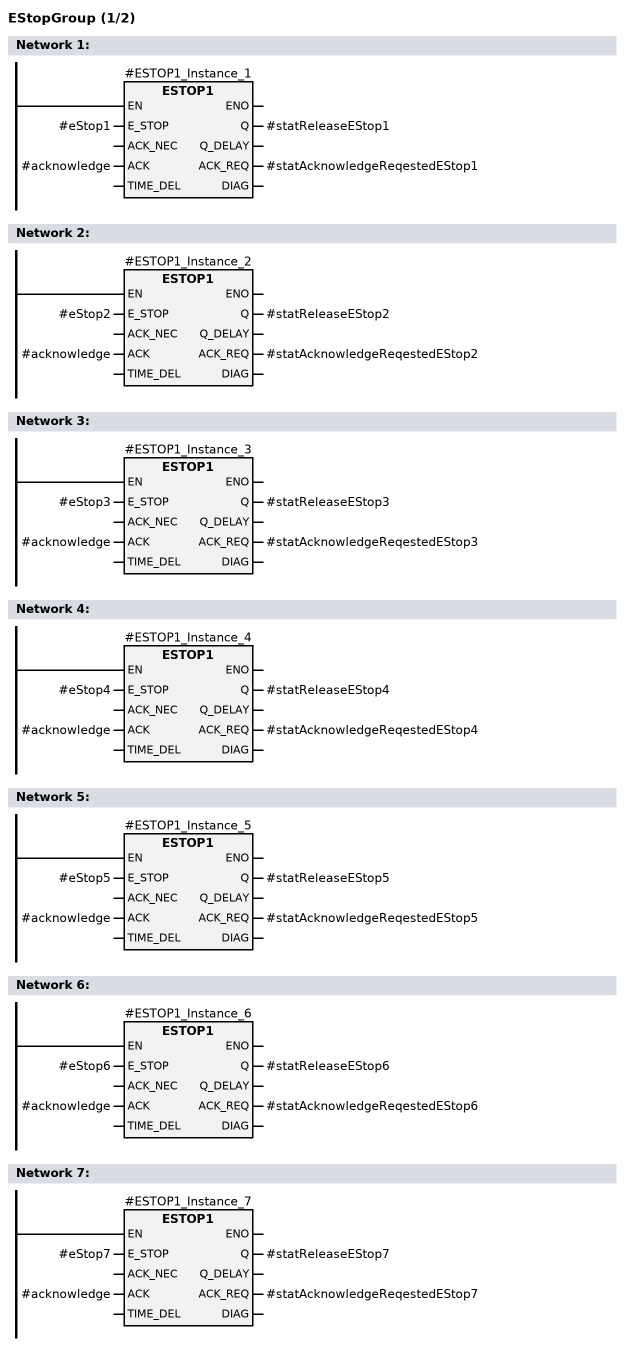
   #ESTOP1_Instance_1(E_STOP := #eStop1,   // ESTOP1
                      ACK := #acknowledge,
                      Q => #statReleaseEStop1,
                      ACK_REQ => #statAcknowledgeReqestedEStop1);
END_REGION

REGION Network 2
   #ESTOP1_Instance_2(E_STOP := #eStop2,   // ESTOP1
                      ACK := #acknowledge,
                      Q => #statReleaseEStop2,
                      ACK_REQ => #statAcknowledgeReqestedEStop2);
END_REGION

REGION Network 3
   #ESTOP1_Instance_3(E_STOP := #eStop3,   // ESTOP1
                      ACK := #acknowledge,
                      Q => #statReleaseEStop3,
                      ACK_REQ => #statAcknowledgeReqestedEStop3);
END_REGION

REGION Network 4
   #ESTOP1_Instance_4(E_STOP := #eStop4,   // ESTOP1
                      ACK := #acknowledge,
                      Q => #statReleaseEStop4,
                      ACK_REQ => #statAcknowledgeReqestedEStop4);
END_REGION

REGION Network 5
   #ESTOP1_Instance_5(E_STOP := #eStop5,   // ESTOP1
                      ACK := #acknowledge,
                      Q => #statReleaseEStop5,
                      ACK_REQ => #statAcknowledgeReqestedEStop5);
END_REGION

REGION Network 6
   #ESTOP1_Instance_6(E_STOP := #eStop6,   // ESTOP1
                      ACK := #acknowledge,
                      Q => #statReleaseEStop6,
                      ACK_REQ => #statAcknowledgeReqestedEStop6);
END_REGION

REGION Network 7
   #ESTOP1_Instance_7(E_STOP := #eStop7,   // ESTOP1
                      ACK := #acknowledge,
                      Q => #statReleaseEStop7,
                      ACK_REQ => #statAcknowledgeReqestedEStop7);
END_REGION

REGION Network 8
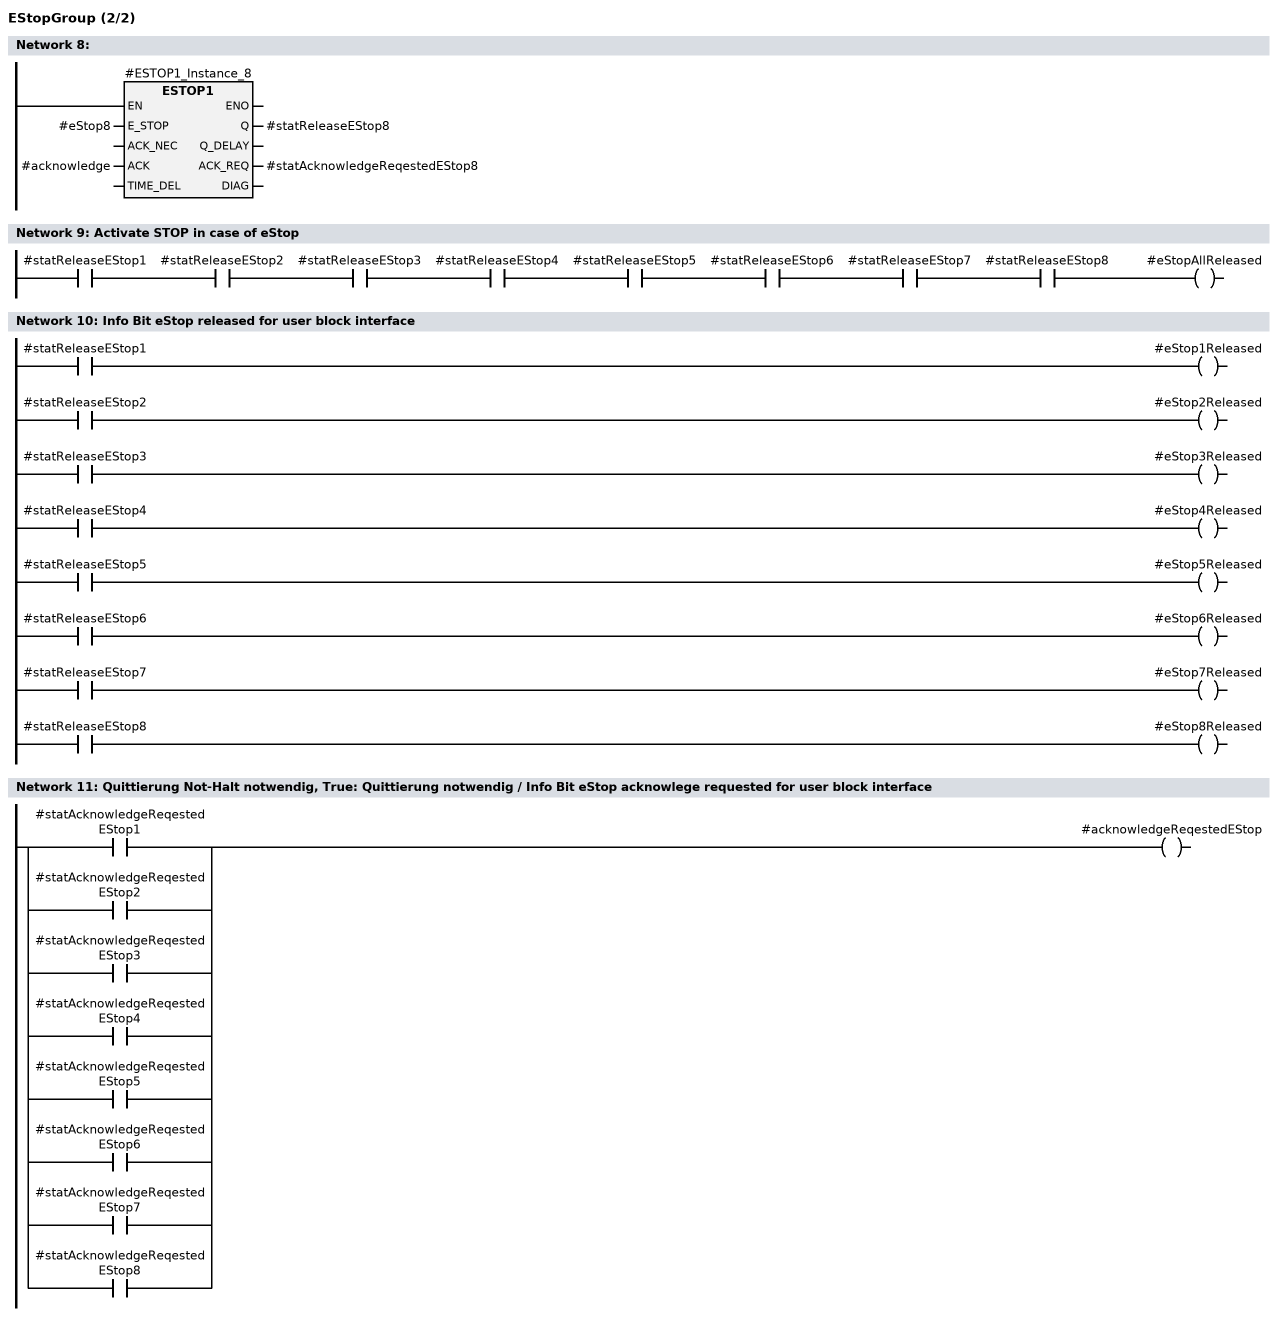
   #ESTOP1_Instance_8(E_STOP := #eStop8,   // ESTOP1
                      ACK := #acknowledge,
                      Q => #statReleaseEStop8,
                      ACK_REQ => #statAcknowledgeReqestedEStop8);
END_REGION

REGION Network 9: Activate STOP in case of eStop
   RUNG wire#powerrail
      Contact( #statReleaseEStop1 )
      Contact( #statReleaseEStop2 )
      Contact( #statReleaseEStop3 )
      Contact( #statReleaseEStop4 )
      Contact( #statReleaseEStop5 )
      Contact( #statReleaseEStop6 )
      Contact( #statReleaseEStop7 )
      Contact( #statReleaseEStop8 )
      Coil( #eStopAllReleased )
   END_RUNG
   // the same network as SCL:
   #eStopAllReleased := #statReleaseEStop1 AND #statReleaseEStop2 AND #statReleaseEStop3 AND #statReleaseEStop4 AND #statReleaseEStop5 AND #statReleaseEStop6 AND #statReleaseEStop7 AND #statReleaseEStop8;
END_REGION

REGION Network 10: Info Bit eStop released for user block interface
   RUNG wire#powerrail
      Contact( #statReleaseEStop1 )
      Coil( #eStop1Released )
   END_RUNG
   RUNG wire#powerrail
      Contact( #statReleaseEStop2 )
      Coil( #eStop2Released )
   END_RUNG
   RUNG wire#powerrail
      Contact( #statReleaseEStop3 )
      Coil( #eStop3Released )
   END_RUNG
   RUNG wire#powerrail
      Contact( #statReleaseEStop4 )
      Coil( #eStop4Released )
   END_RUNG
   RUNG wire#powerrail
      Contact( #statReleaseEStop5 )
      Coil( #eStop5Released )
   END_RUNG
   RUNG wire#powerrail
      Contact( #statReleaseEStop6 )
      Coil( #eStop6Released )
   END_RUNG
   RUNG wire#powerrail
      Contact( #statReleaseEStop7 )
      Coil( #eStop7Released )
   END_RUNG
   RUNG wire#powerrail
      Contact( #statReleaseEStop8 )
      Coil( #eStop8Released )
   END_RUNG
   // the same network as SCL:
   #eStop1Released := #statReleaseEStop1;
   #eStop2Released := #statReleaseEStop2;
   #eStop3Released := #statReleaseEStop3;
   #eStop4Released := #statReleaseEStop4;
   #eStop5Released := #statReleaseEStop5;
   #eStop6Released := #statReleaseEStop6;
   #eStop7Released := #statReleaseEStop7;
   #eStop8Released := #statReleaseEStop8;
END_REGION

REGION Network 11: Quittierung Not-Halt notwendig, True: Quittierung notwendig / Info Bit eStop acknowlege requested for user block interface
   RUNG wire#powerrail
      Contact( #statAcknowledgeReqestedEStop1 )
      wire#w1
      Coil( #acknowledgeReqestedEStop )
   END_RUNG
   RUNG wire#powerrail
      Contact( #statAcknowledgeReqestedEStop2 )
   END_RUNG wire#w1
   RUNG wire#powerrail
      Contact( #statAcknowledgeReqestedEStop3 )
   END_RUNG wire#w1
   RUNG wire#powerrail
      Contact( #statAcknowledgeReqestedEStop4 )
   END_RUNG wire#w1
   RUNG wire#powerrail
      Contact( #statAcknowledgeReqestedEStop5 )
   END_RUNG wire#w1
   RUNG wire#powerrail
      Contact( #statAcknowledgeReqestedEStop6 )
   END_RUNG wire#w1
   RUNG wire#powerrail
      Contact( #statAcknowledgeReqestedEStop7 )
   END_RUNG wire#w1
   RUNG wire#powerrail
      Contact( #statAcknowledgeReqestedEStop8 )
   END_RUNG wire#w1
   // the same network as SCL:
   #acknowledgeReqestedEStop := #statAcknowledgeReqestedEStop1 OR #statAcknowledgeReqestedEStop2 OR #statAcknowledgeReqestedEStop3 OR #statAcknowledgeReqestedEStop4 OR #statAcknowledgeReqestedEStop5 OR #statAcknowledgeReqestedEStop6 OR #statAcknowledgeReqestedEStop7 OR #statAcknowledgeReqestedEStop8;
END_REGION
END_FUNCTION_BLOCK

FUNCTION_BLOCK "LightCurtainGroup"   // FB12, F_LAD
{ S7_Optimized_Access := 'TRUE' }
VERSION : 0.1
   VAR_INPUT
      acknowledge : Bool;   // Acknowledge / Quittierung, Positive Flanke notwendig, NO / Acknowledge, positive signal edge, NO
      selAccZone : Bool;
      entryButtonZone1 : Bool;   // Entry button – Zone 1 (LC 1-6)
      entryButtonZone2 : Bool;   // Entry button – Zone 2 (LC 1, 3, 6)
      entryButtonZone3 : Bool;   // Entry button – Zone 3 (LC 2, 4, 5)
      robotInZone2 : Bool;
      robotInZone3 : Bool;
      lc1Ossd1 : Bool;
      lc1Ossd2 : Bool;
      lc2Ossd1 : Bool;
      lc2Ossd2 : Bool;
      lc3Ossd1 : Bool;
      lc3Ossd2 : Bool;
      lc4Ossd1 : Bool;
      lc4Ossd2 : Bool;
      lc5Ossd1 : Bool;
      lc5Ossd2 : Bool;
      lc6Ossd1 : Bool;
      lc6Ossd2 : Bool;
   END_VAR
   VAR_OUTPUT
      lcAllFree : Bool;   // All light curtains ready
      lc1Free : Bool;   // Light curtain 1 ready
      lc2Free : Bool;
      lc3Free : Bool;   // Light curtain 3 ready
      lc4Free : Bool;
      lc5Free : Bool;
      lc6Free : Bool;   // Light curtain 6 ready
      accessReqZ2 : Bool;
      accessReqZ3 : Bool;
      zone1AccessGranted : Bool;
      zone2AccessGranted : Bool;
      zone3AccessGranted : Bool;
   END_VAR
   VAR
      EV1oo2DI_Instance_1 : EV1oo2DI;
      EV1oo2DI_Instance_2 : EV1oo2DI;
      EV1oo2DI_Instance_3 : EV1oo2DI;
      MUT_P_Instance_1 : MUT_P;
      accZ2Ok : Bool;
      accZ3Ok : Bool;
      lcZone2Free : Bool;
      lcZone3Free : Bool;
      EV1oo2DI_Instance_4 : EV1oo2DI;
      EV1oo2DI_Instance_5 : EV1oo2DI;
      EV1oo2DI_Instance_6 : EV1oo2DI;
   END_VAR
BEGIN

REGION Network 1
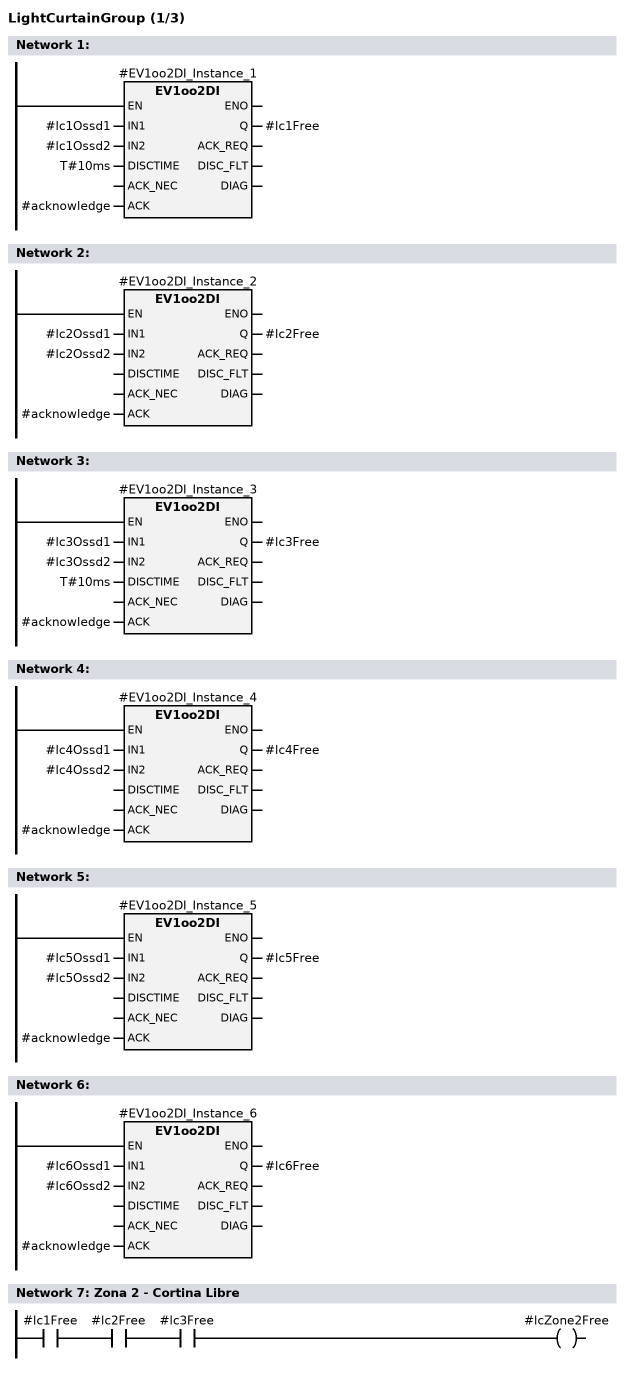
   #EV1oo2DI_Instance_1(IN1 := #lc1Ossd1,   // EV1oo2DI
                        IN2 := #lc1Ossd2,
                        DISCTIME := T#10ms,
                        ACK := #acknowledge,
                        Q => #lc1Free);
END_REGION

REGION Network 2
   #EV1oo2DI_Instance_2(IN1 := #lc2Ossd1, IN2 := #lc2Ossd2, ACK := #acknowledge, Q => #lc2Free);   // EV1oo2DI
END_REGION

REGION Network 3
   #EV1oo2DI_Instance_3(IN1 := #lc3Ossd1,   // EV1oo2DI
                        IN2 := #lc3Ossd2,
                        DISCTIME := T#10ms,
                        ACK := #acknowledge,
                        Q => #lc3Free);
END_REGION

REGION Network 4
   #EV1oo2DI_Instance_4(IN1 := #lc4Ossd1, IN2 := #lc4Ossd2, ACK := #acknowledge, Q => #lc4Free);   // EV1oo2DI
END_REGION

REGION Network 5
   #EV1oo2DI_Instance_5(IN1 := #lc5Ossd1, IN2 := #lc5Ossd2, ACK := #acknowledge, Q => #lc5Free);   // EV1oo2DI
END_REGION

REGION Network 6
   #EV1oo2DI_Instance_6(IN1 := #lc6Ossd1, IN2 := #lc6Ossd2, ACK := #acknowledge, Q => #lc6Free);   // EV1oo2DI
END_REGION

REGION Network 7: Zona 2 - Cortina Libre
   RUNG wire#powerrail
      Contact( #lc1Free )
      Contact( #lc2Free )
      Contact( #lc3Free )
      Coil( #lcZone2Free )
   END_RUNG
   // the same network as SCL:
   #lcZone2Free := #lc1Free AND #lc2Free AND #lc3Free;
END_REGION

REGION Network 8: Zona 3 - Cortina Libre
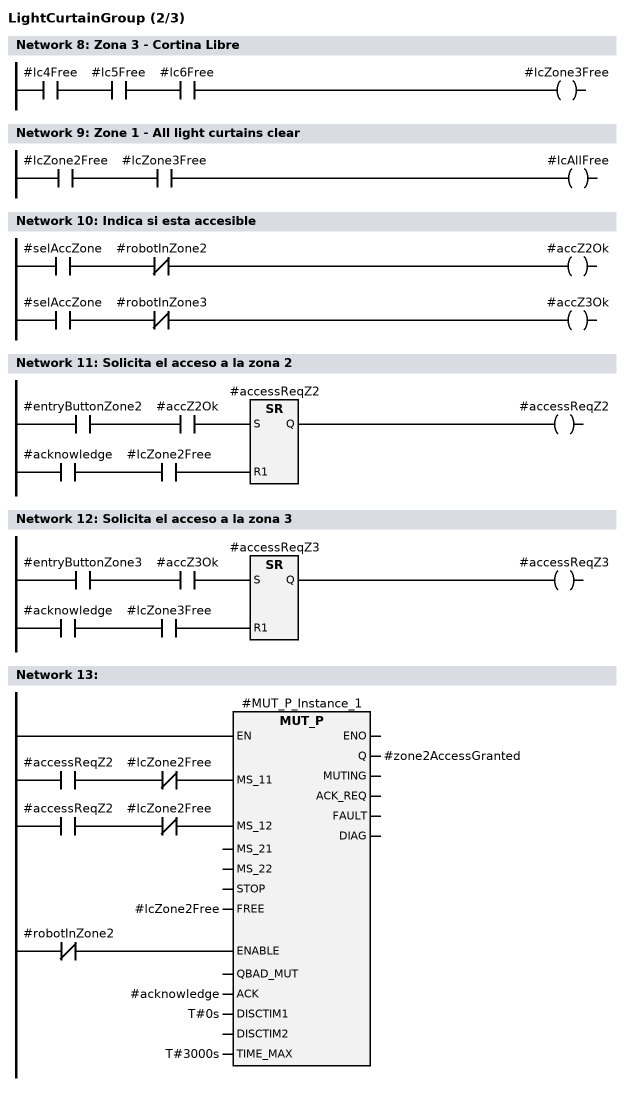
   RUNG wire#powerrail
      Contact( #lc4Free )
      Contact( #lc5Free )
      Contact( #lc6Free )
      Coil( #lcZone3Free )
   END_RUNG
   // the same network as SCL:
   #lcZone3Free := #lc4Free AND #lc5Free AND #lc6Free;
END_REGION

REGION Network 9: Zone 1 - All light curtains clear
   RUNG wire#powerrail
      Contact( #lcZone2Free )
      Contact( #lcZone3Free )
      Coil( #lcAllFree )
   END_RUNG
   // the same network as SCL:
   #lcAllFree := #lcZone2Free AND #lcZone3Free;
END_REGION

REGION Network 10: Indica si esta accesible
   RUNG wire#powerrail
      Contact( #selAccZone )
      I_Contact( #robotInZone2 )
      Coil( #accZ2Ok )
   END_RUNG
   RUNG wire#powerrail
      Contact( #selAccZone )
      I_Contact( #robotInZone3 )
      Coil( #accZ3Ok )
   END_RUNG
   // the same network as SCL:
   #accZ2Ok := #selAccZone AND NOT #robotInZone2;
   #accZ3Ok := #selAccZone AND NOT #robotInZone3;
END_REGION

REGION Network 11: Solicita el acceso a la zona 2
   RUNG wire#powerrail
      Contact( #entryButtonZone2 )
      Contact( #accZ2Ok )
      S_SR(operand := #accessReqZ2, r1 := wire#w1)
      Coil( #accessReqZ2 )
   END_RUNG
   RUNG wire#powerrail
      Contact( #acknowledge )
      Contact( #lcZone2Free )
   END_RUNG wire#w1
   // the same network as SCL:
   IF #entryButtonZone2 AND #accZ2Ok THEN
       #accessReqZ2 := TRUE;   // SR flip-flop
   END_IF;
   IF #acknowledge AND #lcZone2Free THEN #accessReqZ2 := FALSE; END_IF;
   #accessReqZ2 := #accessReqZ2;
END_REGION

REGION Network 12: Solicita el acceso a la zona 3
   RUNG wire#powerrail
      Contact( #entryButtonZone3 )
      Contact( #accZ3Ok )
      S_SR(operand := #accessReqZ3, r1 := wire#w1)
      Coil( #accessReqZ3 )
   END_RUNG
   RUNG wire#powerrail
      Contact( #acknowledge )
      Contact( #lcZone3Free )
   END_RUNG wire#w1
   // the same network as SCL:
   IF #entryButtonZone3 AND #accZ3Ok THEN
       #accessReqZ3 := TRUE;   // SR flip-flop
   END_IF;
   IF #acknowledge AND #lcZone3Free THEN #accessReqZ3 := FALSE; END_IF;
   #accessReqZ3 := #accessReqZ3;
END_REGION

REGION Network 13
   #MUT_P_Instance_1(MS_11 := #accessReqZ2 AND NOT #lcZone2Free,   // MUT_P
                     MS_12 := #accessReqZ2 AND NOT #lcZone2Free,
                     FREE := #lcZone2Free,
                     ENABLE := NOT #robotInZone2,
                     ACK := #acknowledge,
                     DISCTIM1 := T#0s,
                     TIME_MAX := T#3000s,
                     Q => #zone2AccessGranted);
END_REGION

REGION Network 14
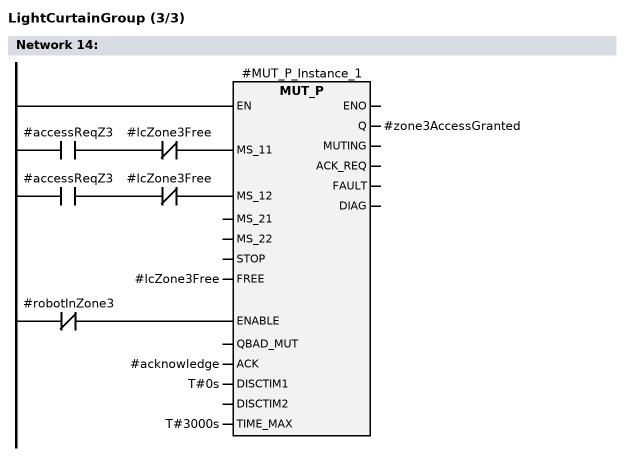
   #MUT_P_Instance_1(MS_11 := #accessReqZ3 AND NOT #lcZone3Free,   // MUT_P
                     MS_12 := #accessReqZ3 AND NOT #lcZone3Free,
                     FREE := #lcZone3Free,
                     ENABLE := NOT #robotInZone3,
                     ACK := #acknowledge,
                     DISCTIM1 := T#0s,
                     TIME_MAX := T#3000s,
                     Q => #zone3AccessGranted);
END_REGION
END_FUNCTION_BLOCK

FUNCTION_BLOCK "SafetyDoor"   // FB13, F_FBD
{ S7_Optimized_Access := 'TRUE' }
VERSION : 0.1
   VAR_OUTPUT
      SAF_DOOR_CLSD_RDY : Bool;   // Safety door closed & locked – ready
   END_VAR
   VAR
      SFDOOR_Instance_1 : SFDOOR;
   END_VAR
BEGIN

REGION Network 1
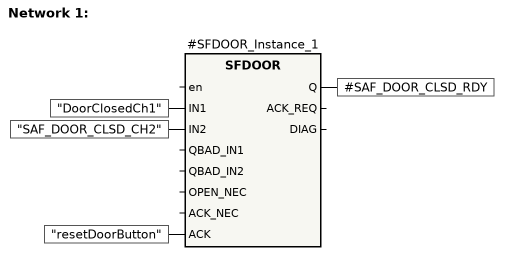
   #SFDOOR_Instance_1(IN1 := "DoorClosedCh1",   // SFDOOR
                      IN2 := "SAF_DOOR_CLSD_CH2",
                      ACK := "resetDoorButton",
                      Q => #SAF_DOOR_CLSD_RDY);
END_REGION
END_FUNCTION_BLOCK

// folder: 410. Festo cuba

FUNCTION_BLOCK "HMI_CUBA"   // FB7, LAD
{ S7_Optimized_Access := 'TRUE' }
VERSION : 0.1
BEGIN

REGION Network 1
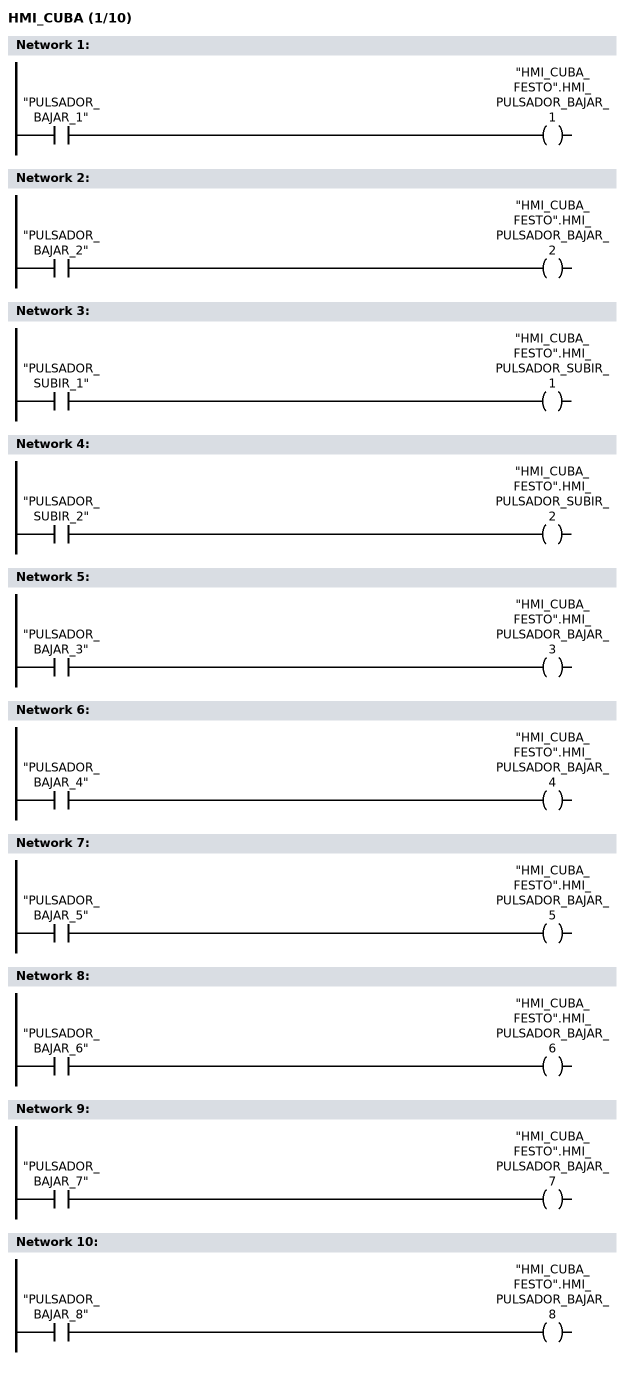
   RUNG wire#powerrail
      Contact( "PULSADOR_BAJAR_1" )
      Coil( "HMI_CUBA_FESTO".HMI_PULSADOR_BAJAR_1 )
   END_RUNG
   // the same network as SCL:
   "HMI_CUBA_FESTO".HMI_PULSADOR_BAJAR_1 := "PULSADOR_BAJAR_1";
END_REGION

REGION Network 2
   RUNG wire#powerrail
      Contact( "PULSADOR_BAJAR_2" )
      Coil( "HMI_CUBA_FESTO".HMI_PULSADOR_BAJAR_2 )
   END_RUNG
   // the same network as SCL:
   "HMI_CUBA_FESTO".HMI_PULSADOR_BAJAR_2 := "PULSADOR_BAJAR_2";
END_REGION

REGION Network 3
   RUNG wire#powerrail
      Contact( "PULSADOR_SUBIR_1" )
      Coil( "HMI_CUBA_FESTO".HMI_PULSADOR_SUBIR_1 )
   END_RUNG
   // the same network as SCL:
   "HMI_CUBA_FESTO".HMI_PULSADOR_SUBIR_1 := "PULSADOR_SUBIR_1";
END_REGION

REGION Network 4
   RUNG wire#powerrail
      Contact( "PULSADOR_SUBIR_2" )
      Coil( "HMI_CUBA_FESTO".HMI_PULSADOR_SUBIR_2 )
   END_RUNG
   // the same network as SCL:
   "HMI_CUBA_FESTO".HMI_PULSADOR_SUBIR_2 := "PULSADOR_SUBIR_2";
END_REGION

REGION Network 5
   RUNG wire#powerrail
      Contact( "PULSADOR_BAJAR_3" )
      Coil( "HMI_CUBA_FESTO".HMI_PULSADOR_BAJAR_3 )
   END_RUNG
   // the same network as SCL:
   "HMI_CUBA_FESTO".HMI_PULSADOR_BAJAR_3 := "PULSADOR_BAJAR_3";
END_REGION

REGION Network 6
   RUNG wire#powerrail
      Contact( "PULSADOR_BAJAR_4" )
      Coil( "HMI_CUBA_FESTO".HMI_PULSADOR_BAJAR_4 )
   END_RUNG
   // the same network as SCL:
   "HMI_CUBA_FESTO".HMI_PULSADOR_BAJAR_4 := "PULSADOR_BAJAR_4";
END_REGION

REGION Network 7
   RUNG wire#powerrail
      Contact( "PULSADOR_BAJAR_5" )
      Coil( "HMI_CUBA_FESTO".HMI_PULSADOR_BAJAR_5 )
   END_RUNG
   // the same network as SCL:
   "HMI_CUBA_FESTO".HMI_PULSADOR_BAJAR_5 := "PULSADOR_BAJAR_5";
END_REGION

REGION Network 8
   RUNG wire#powerrail
      Contact( "PULSADOR_BAJAR_6" )
      Coil( "HMI_CUBA_FESTO".HMI_PULSADOR_BAJAR_6 )
   END_RUNG
   // the same network as SCL:
   "HMI_CUBA_FESTO".HMI_PULSADOR_BAJAR_6 := "PULSADOR_BAJAR_6";
END_REGION

REGION Network 9
   RUNG wire#powerrail
      Contact( "PULSADOR_BAJAR_7" )
      Coil( "HMI_CUBA_FESTO".HMI_PULSADOR_BAJAR_7 )
   END_RUNG
   // the same network as SCL:
   "HMI_CUBA_FESTO".HMI_PULSADOR_BAJAR_7 := "PULSADOR_BAJAR_7";
END_REGION

REGION Network 10
   RUNG wire#powerrail
      Contact( "PULSADOR_BAJAR_8" )
      Coil( "HMI_CUBA_FESTO".HMI_PULSADOR_BAJAR_8 )
   END_RUNG
   // the same network as SCL:
   "HMI_CUBA_FESTO".HMI_PULSADOR_BAJAR_8 := "PULSADOR_BAJAR_8";
END_REGION

REGION Network 11
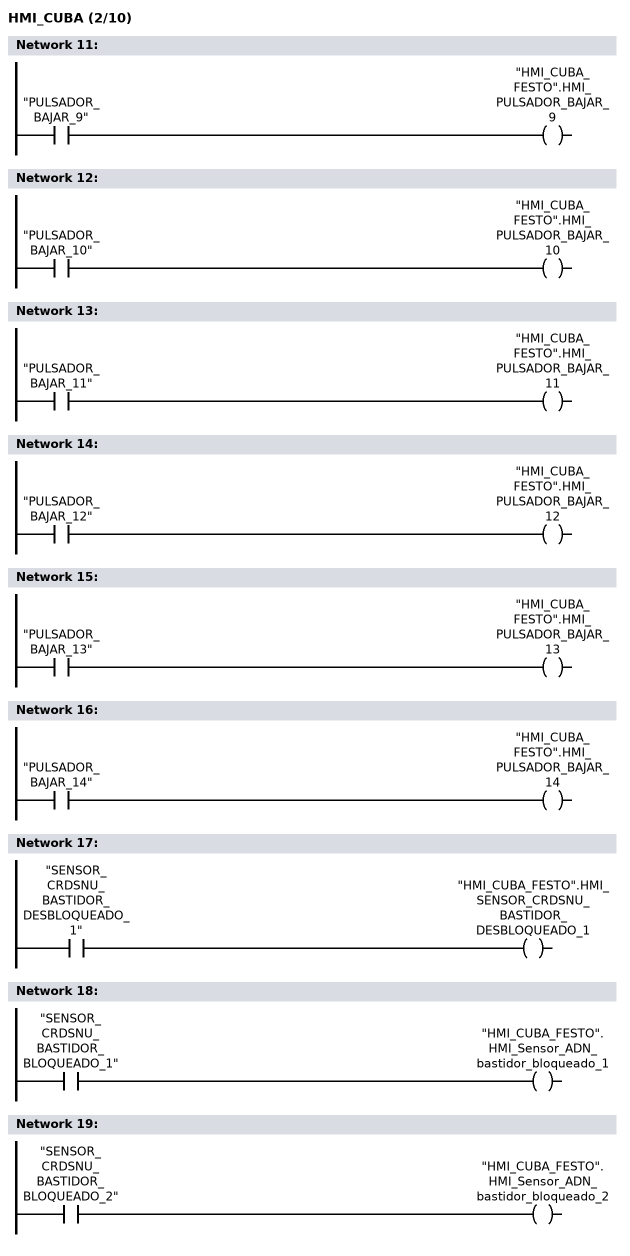
   RUNG wire#powerrail
      Contact( "PULSADOR_BAJAR_9" )
      Coil( "HMI_CUBA_FESTO".HMI_PULSADOR_BAJAR_9 )
   END_RUNG
   // the same network as SCL:
   "HMI_CUBA_FESTO".HMI_PULSADOR_BAJAR_9 := "PULSADOR_BAJAR_9";
END_REGION

REGION Network 12
   RUNG wire#powerrail
      Contact( "PULSADOR_BAJAR_10" )
      Coil( "HMI_CUBA_FESTO".HMI_PULSADOR_BAJAR_10 )
   END_RUNG
   // the same network as SCL:
   "HMI_CUBA_FESTO".HMI_PULSADOR_BAJAR_10 := "PULSADOR_BAJAR_10";
END_REGION

REGION Network 13
   RUNG wire#powerrail
      Contact( "PULSADOR_BAJAR_11" )
      Coil( "HMI_CUBA_FESTO".HMI_PULSADOR_BAJAR_11 )
   END_RUNG
   // the same network as SCL:
   "HMI_CUBA_FESTO".HMI_PULSADOR_BAJAR_11 := "PULSADOR_BAJAR_11";
END_REGION

REGION Network 14
   RUNG wire#powerrail
      Contact( "PULSADOR_BAJAR_12" )
      Coil( "HMI_CUBA_FESTO".HMI_PULSADOR_BAJAR_12 )
   END_RUNG
   // the same network as SCL:
   "HMI_CUBA_FESTO".HMI_PULSADOR_BAJAR_12 := "PULSADOR_BAJAR_12";
END_REGION

REGION Network 15
   RUNG wire#powerrail
      Contact( "PULSADOR_BAJAR_13" )
      Coil( "HMI_CUBA_FESTO".HMI_PULSADOR_BAJAR_13 )
   END_RUNG
   // the same network as SCL:
   "HMI_CUBA_FESTO".HMI_PULSADOR_BAJAR_13 := "PULSADOR_BAJAR_13";
END_REGION

REGION Network 16
   RUNG wire#powerrail
      Contact( "PULSADOR_BAJAR_14" )
      Coil( "HMI_CUBA_FESTO".HMI_PULSADOR_BAJAR_14 )
   END_RUNG
   // the same network as SCL:
   "HMI_CUBA_FESTO".HMI_PULSADOR_BAJAR_14 := "PULSADOR_BAJAR_14";
END_REGION

REGION Network 17
   RUNG wire#powerrail
      Contact( "SENSOR_CRDSNU_BASTIDOR_DESBLOQUEADO_1" )
      Coil( "HMI_CUBA_FESTO".HMI_SENSOR_CRDSNU_BASTIDOR_DESBLOQUEADO_1 )
   END_RUNG
   // the same network as SCL:
   "HMI_CUBA_FESTO".HMI_SENSOR_CRDSNU_BASTIDOR_DESBLOQUEADO_1 := "SENSOR_CRDSNU_BASTIDOR_DESBLOQUEADO_1";
END_REGION

REGION Network 18
   RUNG wire#powerrail
      Contact( "SENSOR_CRDSNU_BASTIDOR_BLOQUEADO_1" )
      Coil( "HMI_CUBA_FESTO".HMI_Sensor_ADN_bastidor_bloqueado_1 )
   END_RUNG
   // the same network as SCL:
   "HMI_CUBA_FESTO".HMI_Sensor_ADN_bastidor_bloqueado_1 := "SENSOR_CRDSNU_BASTIDOR_BLOQUEADO_1";
END_REGION

REGION Network 19
   RUNG wire#powerrail
      Contact( "SENSOR_CRDSNU_BASTIDOR_BLOQUEADO_2" )
      Coil( "HMI_CUBA_FESTO".HMI_Sensor_ADN_bastidor_bloqueado_2 )
   END_RUNG
   // the same network as SCL:
   "HMI_CUBA_FESTO".HMI_Sensor_ADN_bastidor_bloqueado_2 := "SENSOR_CRDSNU_BASTIDOR_BLOQUEADO_2";
END_REGION

REGION Network 20
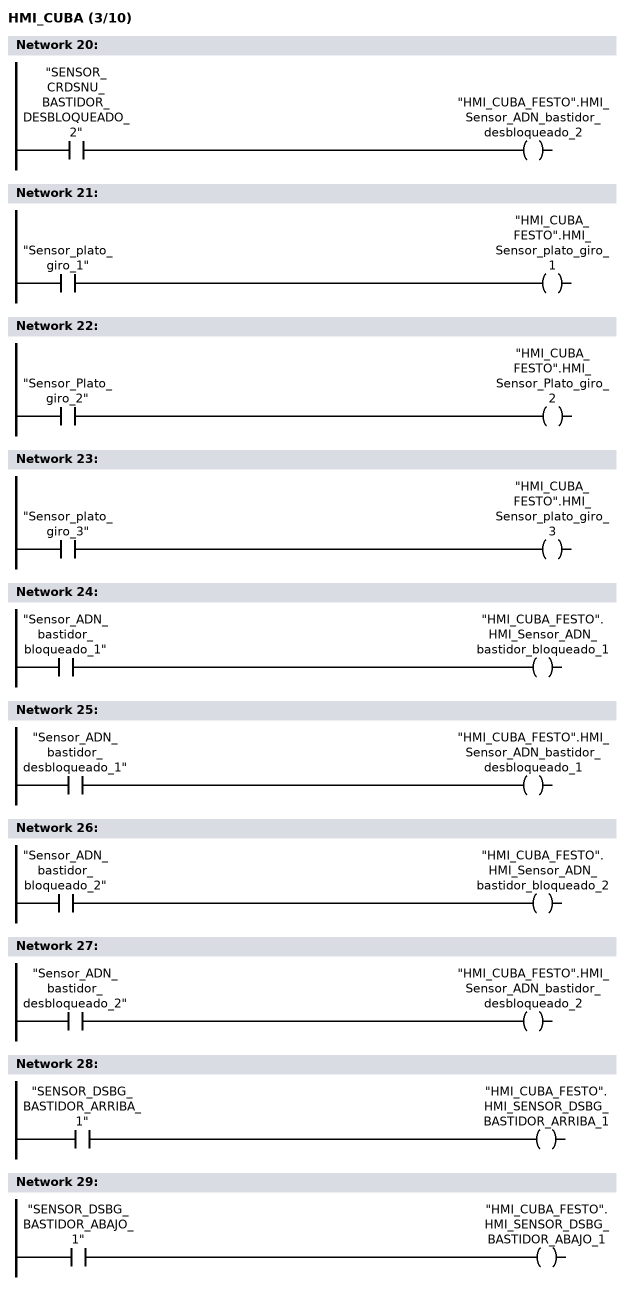
   RUNG wire#powerrail
      Contact( "SENSOR_CRDSNU_BASTIDOR_DESBLOQUEADO_2" )
      Coil( "HMI_CUBA_FESTO".HMI_Sensor_ADN_bastidor_desbloqueado_2 )
   END_RUNG
   // the same network as SCL:
   "HMI_CUBA_FESTO".HMI_Sensor_ADN_bastidor_desbloqueado_2 := "SENSOR_CRDSNU_BASTIDOR_DESBLOQUEADO_2";
END_REGION

REGION Network 21
   RUNG wire#powerrail
      Contact( "Sensor_plato_giro_1" )
      Coil( "HMI_CUBA_FESTO".HMI_Sensor_plato_giro_1 )
   END_RUNG
   // the same network as SCL:
   "HMI_CUBA_FESTO".HMI_Sensor_plato_giro_1 := "Sensor_plato_giro_1";
END_REGION

REGION Network 22
   RUNG wire#powerrail
      Contact( "Sensor_Plato_giro_2" )
      Coil( "HMI_CUBA_FESTO".HMI_Sensor_Plato_giro_2 )
   END_RUNG
   // the same network as SCL:
   "HMI_CUBA_FESTO".HMI_Sensor_Plato_giro_2 := "Sensor_Plato_giro_2";
END_REGION

REGION Network 23
   RUNG wire#powerrail
      Contact( "Sensor_plato_giro_3" )
      Coil( "HMI_CUBA_FESTO".HMI_Sensor_plato_giro_3 )
   END_RUNG
   // the same network as SCL:
   "HMI_CUBA_FESTO".HMI_Sensor_plato_giro_3 := "Sensor_plato_giro_3";
END_REGION

REGION Network 24
   RUNG wire#powerrail
      Contact( "Sensor_ADN_bastidor_bloqueado_1" )
      Coil( "HMI_CUBA_FESTO".HMI_Sensor_ADN_bastidor_bloqueado_1 )
   END_RUNG
   // the same network as SCL:
   "HMI_CUBA_FESTO".HMI_Sensor_ADN_bastidor_bloqueado_1 := "Sensor_ADN_bastidor_bloqueado_1";
END_REGION

REGION Network 25
   RUNG wire#powerrail
      Contact( "Sensor_ADN_bastidor_desbloqueado_1" )
      Coil( "HMI_CUBA_FESTO".HMI_Sensor_ADN_bastidor_desbloqueado_1 )
   END_RUNG
   // the same network as SCL:
   "HMI_CUBA_FESTO".HMI_Sensor_ADN_bastidor_desbloqueado_1 := "Sensor_ADN_bastidor_desbloqueado_1";
END_REGION

REGION Network 26
   RUNG wire#powerrail
      Contact( "Sensor_ADN_bastidor_bloqueado_2" )
      Coil( "HMI_CUBA_FESTO".HMI_Sensor_ADN_bastidor_bloqueado_2 )
   END_RUNG
   // the same network as SCL:
   "HMI_CUBA_FESTO".HMI_Sensor_ADN_bastidor_bloqueado_2 := "Sensor_ADN_bastidor_bloqueado_2";
END_REGION

REGION Network 27
   RUNG wire#powerrail
      Contact( "Sensor_ADN_bastidor_desbloqueado_2" )
      Coil( "HMI_CUBA_FESTO".HMI_Sensor_ADN_bastidor_desbloqueado_2 )
   END_RUNG
   // the same network as SCL:
   "HMI_CUBA_FESTO".HMI_Sensor_ADN_bastidor_desbloqueado_2 := "Sensor_ADN_bastidor_desbloqueado_2";
END_REGION

REGION Network 28
   RUNG wire#powerrail
      Contact( "SENSOR_DSBG_BASTIDOR_ARRIBA_1" )
      Coil( "HMI_CUBA_FESTO".HMI_SENSOR_DSBG_BASTIDOR_ARRIBA_1 )
   END_RUNG
   // the same network as SCL:
   "HMI_CUBA_FESTO".HMI_SENSOR_DSBG_BASTIDOR_ARRIBA_1 := "SENSOR_DSBG_BASTIDOR_ARRIBA_1";
END_REGION

REGION Network 29
   RUNG wire#powerrail
      Contact( "SENSOR_DSBG_BASTIDOR_ABAJO_1" )
      Coil( "HMI_CUBA_FESTO".HMI_SENSOR_DSBG_BASTIDOR_ABAJO_1 )
   END_RUNG
   // the same network as SCL:
   "HMI_CUBA_FESTO".HMI_SENSOR_DSBG_BASTIDOR_ABAJO_1 := "SENSOR_DSBG_BASTIDOR_ABAJO_1";
END_REGION

REGION Network 30
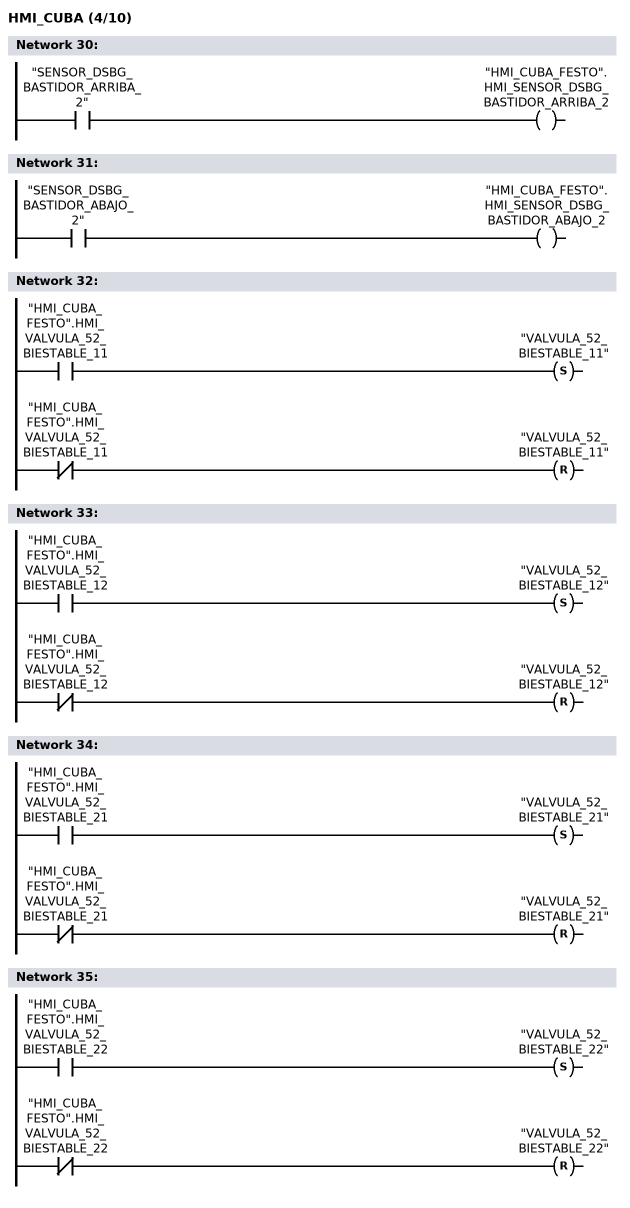
   RUNG wire#powerrail
      Contact( "SENSOR_DSBG_BASTIDOR_ARRIBA_2" )
      Coil( "HMI_CUBA_FESTO".HMI_SENSOR_DSBG_BASTIDOR_ARRIBA_2 )
   END_RUNG
   // the same network as SCL:
   "HMI_CUBA_FESTO".HMI_SENSOR_DSBG_BASTIDOR_ARRIBA_2 := "SENSOR_DSBG_BASTIDOR_ARRIBA_2";
END_REGION

REGION Network 31
   RUNG wire#powerrail
      Contact( "SENSOR_DSBG_BASTIDOR_ABAJO_2" )
      Coil( "HMI_CUBA_FESTO".HMI_SENSOR_DSBG_BASTIDOR_ABAJO_2 )
   END_RUNG
   // the same network as SCL:
   "HMI_CUBA_FESTO".HMI_SENSOR_DSBG_BASTIDOR_ABAJO_2 := "SENSOR_DSBG_BASTIDOR_ABAJO_2";
END_REGION

REGION Network 32
   RUNG wire#powerrail
      Contact( "HMI_CUBA_FESTO".HMI_VALVULA_52_BIESTABLE_11 )
      S_Coil( "VALVULA_52_BIESTABLE_11" )
   END_RUNG
   RUNG wire#powerrail
      I_Contact( "HMI_CUBA_FESTO".HMI_VALVULA_52_BIESTABLE_11 )
      R_Coil( "VALVULA_52_BIESTABLE_11" )
   END_RUNG
   // the same network as SCL:
   IF "HMI_CUBA_FESTO".HMI_VALVULA_52_BIESTABLE_11 THEN "VALVULA_52_BIESTABLE_11" := TRUE; END_IF;
   IF NOT "HMI_CUBA_FESTO".HMI_VALVULA_52_BIESTABLE_11 THEN "VALVULA_52_BIESTABLE_11" := FALSE; END_IF;
END_REGION

REGION Network 33
   RUNG wire#powerrail
      Contact( "HMI_CUBA_FESTO".HMI_VALVULA_52_BIESTABLE_12 )
      S_Coil( "VALVULA_52_BIESTABLE_12" )
   END_RUNG
   RUNG wire#powerrail
      I_Contact( "HMI_CUBA_FESTO".HMI_VALVULA_52_BIESTABLE_12 )
      R_Coil( "VALVULA_52_BIESTABLE_12" )
   END_RUNG
   // the same network as SCL:
   IF "HMI_CUBA_FESTO".HMI_VALVULA_52_BIESTABLE_12 THEN "VALVULA_52_BIESTABLE_12" := TRUE; END_IF;
   IF NOT "HMI_CUBA_FESTO".HMI_VALVULA_52_BIESTABLE_12 THEN "VALVULA_52_BIESTABLE_12" := FALSE; END_IF;
END_REGION

REGION Network 34
   RUNG wire#powerrail
      Contact( "HMI_CUBA_FESTO".HMI_VALVULA_52_BIESTABLE_21 )
      S_Coil( "VALVULA_52_BIESTABLE_21" )
   END_RUNG
   RUNG wire#powerrail
      I_Contact( "HMI_CUBA_FESTO".HMI_VALVULA_52_BIESTABLE_21 )
      R_Coil( "VALVULA_52_BIESTABLE_21" )
   END_RUNG
   // the same network as SCL:
   IF "HMI_CUBA_FESTO".HMI_VALVULA_52_BIESTABLE_21 THEN "VALVULA_52_BIESTABLE_21" := TRUE; END_IF;
   IF NOT "HMI_CUBA_FESTO".HMI_VALVULA_52_BIESTABLE_21 THEN "VALVULA_52_BIESTABLE_21" := FALSE; END_IF;
END_REGION

REGION Network 35
   RUNG wire#powerrail
      Contact( "HMI_CUBA_FESTO".HMI_VALVULA_52_BIESTABLE_22 )
      S_Coil( "VALVULA_52_BIESTABLE_22" )
   END_RUNG
   RUNG wire#powerrail
      I_Contact( "HMI_CUBA_FESTO".HMI_VALVULA_52_BIESTABLE_22 )
      R_Coil( "VALVULA_52_BIESTABLE_22" )
   END_RUNG
   // the same network as SCL:
   IF "HMI_CUBA_FESTO".HMI_VALVULA_52_BIESTABLE_22 THEN "VALVULA_52_BIESTABLE_22" := TRUE; END_IF;
   IF NOT "HMI_CUBA_FESTO".HMI_VALVULA_52_BIESTABLE_22 THEN "VALVULA_52_BIESTABLE_22" := FALSE; END_IF;
END_REGION

REGION Network 36
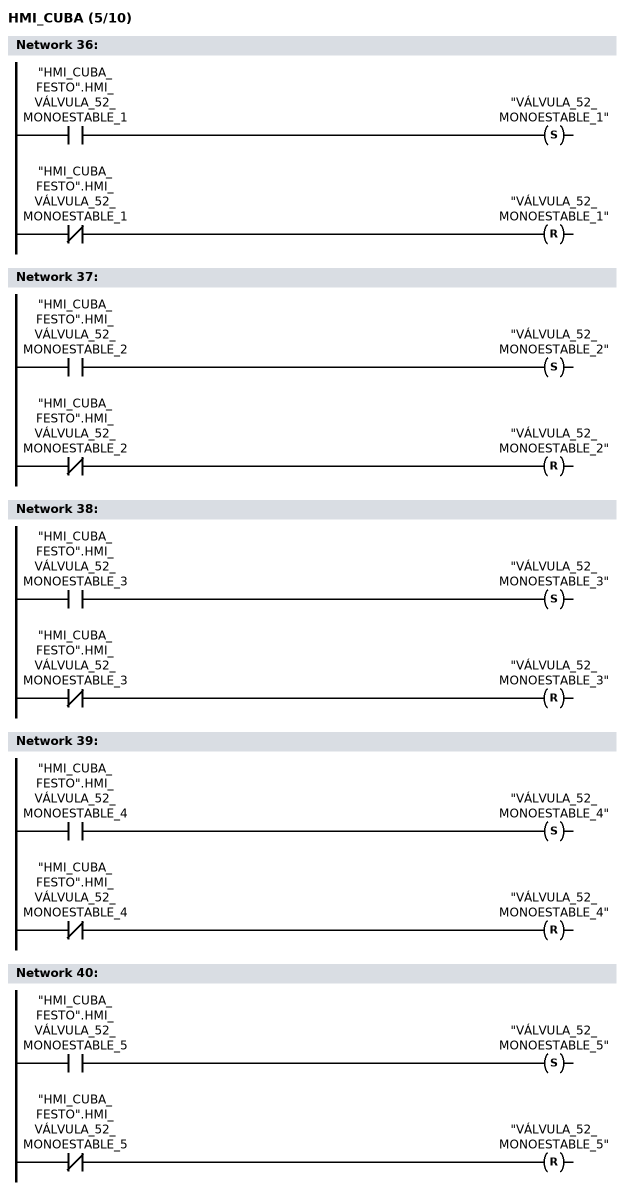
   RUNG wire#powerrail
      Contact( "HMI_CUBA_FESTO".HMI_VÁLVULA_52_MONOESTABLE_1 )
      S_Coil( "VÁLVULA_52_MONOESTABLE_1" )
   END_RUNG
   RUNG wire#powerrail
      I_Contact( "HMI_CUBA_FESTO".HMI_VÁLVULA_52_MONOESTABLE_1 )
      R_Coil( "VÁLVULA_52_MONOESTABLE_1" )
   END_RUNG
   // the same network as SCL:
   IF "HMI_CUBA_FESTO".HMI_VÁLVULA_52_MONOESTABLE_1 THEN "VÁLVULA_52_MONOESTABLE_1" := TRUE; END_IF;
   IF NOT "HMI_CUBA_FESTO".HMI_VÁLVULA_52_MONOESTABLE_1 THEN "VÁLVULA_52_MONOESTABLE_1" := FALSE; END_IF;
END_REGION

REGION Network 37
   RUNG wire#powerrail
      Contact( "HMI_CUBA_FESTO".HMI_VÁLVULA_52_MONOESTABLE_2 )
      S_Coil( "VÁLVULA_52_MONOESTABLE_2" )
   END_RUNG
   RUNG wire#powerrail
      I_Contact( "HMI_CUBA_FESTO".HMI_VÁLVULA_52_MONOESTABLE_2 )
      R_Coil( "VÁLVULA_52_MONOESTABLE_2" )
   END_RUNG
   // the same network as SCL:
   IF "HMI_CUBA_FESTO".HMI_VÁLVULA_52_MONOESTABLE_2 THEN "VÁLVULA_52_MONOESTABLE_2" := TRUE; END_IF;
   IF NOT "HMI_CUBA_FESTO".HMI_VÁLVULA_52_MONOESTABLE_2 THEN "VÁLVULA_52_MONOESTABLE_2" := FALSE; END_IF;
END_REGION

REGION Network 38
   RUNG wire#powerrail
      Contact( "HMI_CUBA_FESTO".HMI_VÁLVULA_52_MONOESTABLE_3 )
      S_Coil( "VÁLVULA_52_MONOESTABLE_3" )
   END_RUNG
   RUNG wire#powerrail
      I_Contact( "HMI_CUBA_FESTO".HMI_VÁLVULA_52_MONOESTABLE_3 )
      R_Coil( "VÁLVULA_52_MONOESTABLE_3" )
   END_RUNG
   // the same network as SCL:
   IF "HMI_CUBA_FESTO".HMI_VÁLVULA_52_MONOESTABLE_3 THEN "VÁLVULA_52_MONOESTABLE_3" := TRUE; END_IF;
   IF NOT "HMI_CUBA_FESTO".HMI_VÁLVULA_52_MONOESTABLE_3 THEN "VÁLVULA_52_MONOESTABLE_3" := FALSE; END_IF;
END_REGION

